(* Logix 5000 project; controller UOWHF Emulate 5570 rev 30.12; software revision 30.00; part 8 of 13 *)
(* tags used below, declared in another part *)
   UOWHF_Add_c : DINT;
   UOWHF_Msg : DINT[16];
   UOWHF_Result : DINT[16];
(* MainProgram, continued *)

   		UOWHF_Result[7]:=UOWHF_Result[7] + 421348795+UOWHF_Add_c;
   		UOWHF_Add_c.7:=UOWHF_Result[7].31;
   		UOWHF_Result[7].31:=0;
   		UOWHF_Result[8]:=UOWHF_Result[8] + 1440025142+UOWHF_Add_c;
   		UOWHF_Add_c.8:=UOWHF_Result[8].31;
   		UOWHF_Result[8].31:=0;
   	End_If;
   	If UOWHF_Msg[2].[17] Then
   		UOWHF_Result[0]:=UOWHF_Result[0] + 1919227168+UOWHF_Add_c;
   		UOWHF_Add_c.0:=UOWHF_Result[0].31;
   		UOWHF_Result[0].31:=0;
   		UOWHF_Result[1]:=UOWHF_Result[1] + 29463341+UOWHF_Add_c;
   		UOWHF_Add_c.1:=UOWHF_Result[1].31;
   		UOWHF_Result[1].31:=0;
   		UOWHF_Result[2]:=UOWHF_Result[2] + 852012451+UOWHF_Add_c;
   		UOWHF_Add_c.2:=UOWHF_Result[2].31;
   		UOWHF_Result[2].31:=0;
   		UOWHF_Result[3]:=UOWHF_Result[3] + 551239594+UOWHF_Add_c;
   		UOWHF_Add_c.3:=UOWHF_Result[3].31;
   		UOWHF_Result[3].31:=0;
   		UOWHF_Result[4]:=UOWHF_Result[4] + 213735753+UOWHF_Add_c;
   		UOWHF_Add_c.4:=UOWHF_Result[4].31;
   		UOWHF_Result[4].31:=0;
   		UOWHF_Result[5]:=UOWHF_Result[5] + 930229489+UOWHF_Add_c;
   		UOWHF_Add_c.5:=UOWHF_Result[5].31;
   		UOWHF_Result[5].31:=0;
   		UOWHF_Result[6]:=UOWHF_Result[6] + 403306511+UOWHF_Add_c;
   		UOWHF_Add_c.6:=UOWHF_Result[6].31;
   		UOWHF_Result[6].31:=0;
   		UOWHF_Result[7]:=UOWHF_Result[7] + 1320163597+UOWHF_Add_c;
   		UOWHF_Add_c.7:=UOWHF_Result[7].31;
   		UOWHF_Result[7].31:=0;
   		UOWHF_Result[8]:=UOWHF_Result[8] + 1897862563+UOWHF_Add_c;
   		UOWHF_Add_c.8:=UOWHF_Result[8].31;
   		UOWHF_Result[8].31:=0;
   	End_If;
   	If UOWHF_Msg[2].[18] Then
   		UOWHF_Result[0]:=UOWHF_Result[0] + 207957642+UOWHF_Add_c;
   		UOWHF_Add_c.0:=UOWHF_Result[0].31;
   		UOWHF_Result[0].31:=0;
   		UOWHF_Result[1]:=UOWHF_Result[1] + 1171801270+UOWHF_Add_c;
   		UOWHF_Add_c.1:=UOWHF_Result[1].31;
   		UOWHF_Result[1].31:=0;
   		UOWHF_Result[2]:=UOWHF_Result[2] + 490989868+UOWHF_Add_c;
   		UOWHF_Add_c.2:=UOWHF_Result[2].31;
   		UOWHF_Result[2].31:=0;
   		UOWHF_Result[3]:=UOWHF_Result[3] + 517478476+UOWHF_Add_c;
   		UOWHF_Add_c.3:=UOWHF_Result[3].31;
   		UOWHF_Result[3].31:=0;
   		UOWHF_Result[4]:=UOWHF_Result[4] + 709606705+UOWHF_Add_c;
   		UOWHF_Add_c.4:=UOWHF_Result[4].31;
   		UOWHF_Result[4].31:=0;
   		UOWHF_Result[5]:=UOWHF_Result[5] + 959699469+UOWHF_Add_c;
   		UOWHF_Add_c.5:=UOWHF_Result[5].31;
   		UOWHF_Result[5].31:=0;
   		UOWHF_Result[6]:=UOWHF_Result[6] + 1426433136+UOWHF_Add_c;
   		UOWHF_Add_c.6:=UOWHF_Result[6].31;
   		UOWHF_Result[6].31:=0;
   		UOWHF_Result[7]:=UOWHF_Result[7] + 861500679+UOWHF_Add_c;
   		UOWHF_Add_c.7:=UOWHF_Result[7].31;
   		UOWHF_Result[7].31:=0;
   		UOWHF_Result[8]:=UOWHF_Result[8] + 1202438537+UOWHF_Add_c;
   		UOWHF_Add_c.8:=UOWHF_Result[8].31;
   		UOWHF_Result[8].31:=0;
   	End_If;
   	If UOWHF_Msg[2].[19] Then
   		UOWHF_Result[0]:=UOWHF_Result[0] + 1004597840+UOWHF_Add_c;
   		UOWHF_Add_c.0:=UOWHF_Result[0].31;
   		UOWHF_Result[0].31:=0;
   		UOWHF_Result[1]:=UOWHF_Result[1] + 599270858+UOWHF_Add_c;
   		UOWHF_Add_c.1:=UOWHF_Result[1].31;
   		UOWHF_Result[1].31:=0;
   		UOWHF_Result[2]:=UOWHF_Result[2] + 334847739+UOWHF_Add_c;
   		UOWHF_Add_c.2:=UOWHF_Result[2].31;
   		UOWHF_Result[2].31:=0;
   		UOWHF_Result[3]:=UOWHF_Result[3] + 1969220087+UOWHF_Add_c;
   		UOWHF_Add_c.3:=UOWHF_Result[3].31;
   		UOWHF_Result[3].31:=0;
   		UOWHF_Result[4]:=UOWHF_Result[4] + 935752387+UOWHF_Add_c;
   		UOWHF_Add_c.4:=UOWHF_Result[4].31;
   		UOWHF_Result[4].31:=0;
   		UOWHF_Result[5]:=UOWHF_Result[5] + 1383478312+UOWHF_Add_c;
   		UOWHF_Add_c.5:=UOWHF_Result[5].31;
   		UOWHF_Result[5].31:=0;
   		UOWHF_Result[6]:=UOWHF_Result[6] + 138334567+UOWHF_Add_c;
   		UOWHF_Add_c.6:=UOWHF_Result[6].31;
   		UOWHF_Result[6].31:=0;
   		UOWHF_Result[7]:=UOWHF_Result[7] + 1365274530+UOWHF_Add_c;
   		UOWHF_Add_c.7:=UOWHF_Result[7].31;
   		UOWHF_Result[7].31:=0;
   		UOWHF_Result[8]:=UOWHF_Result[8] + 534270135+UOWHF_Add_c;
   		UOWHF_Add_c.8:=UOWHF_Result[8].31;
   		UOWHF_Result[8].31:=0;
   	End_If;
   	If UOWHF_Msg[2].[20] Then
   		UOWHF_Result[0]:=UOWHF_Result[0] + 638769264+UOWHF_Add_c;
   		UOWHF_Add_c.0:=UOWHF_Result[0].31;
   		UOWHF_Result[0].31:=0;
   		UOWHF_Result[1]:=UOWHF_Result[1] + 317214964+UOWHF_Add_c;
   		UOWHF_Add_c.1:=UOWHF_Result[1].31;
   		UOWHF_Result[1].31:=0;
   		UOWHF_Result[2]:=UOWHF_Result[2] + 908553039+UOWHF_Add_c;
   		UOWHF_Add_c.2:=UOWHF_Result[2].31;
   		UOWHF_Result[2].31:=0;
   		UOWHF_Result[3]:=UOWHF_Result[3] + 1054049644+UOWHF_Add_c;
   		UOWHF_Add_c.3:=UOWHF_Result[3].31;
   		UOWHF_Result[3].31:=0;
   		UOWHF_Result[4]:=UOWHF_Result[4] + 1355262167+UOWHF_Add_c;
   		UOWHF_Add_c.4:=UOWHF_Result[4].31;
   		UOWHF_Result[4].31:=0;
   		UOWHF_Result[5]:=UOWHF_Result[5] + 1333398518+UOWHF_Add_c;
   		UOWHF_Add_c.5:=UOWHF_Result[5].31;
   		UOWHF_Result[5].31:=0;
   		UOWHF_Result[6]:=UOWHF_Result[6] + 923137105+UOWHF_Add_c;
   		UOWHF_Add_c.6:=UOWHF_Result[6].31;
   		UOWHF_Result[6].31:=0;
   		UOWHF_Result[7]:=UOWHF_Result[7] + 1603787279+UOWHF_Add_c;
   		UOWHF_Add_c.7:=UOWHF_Result[7].31;
   		UOWHF_Result[7].31:=0;
   		UOWHF_Result[8]:=UOWHF_Result[8] + 215241896+UOWHF_Add_c;
   		UOWHF_Add_c.8:=UOWHF_Result[8].31;
   		UOWHF_Result[8].31:=0;
   	End_If;
   	If UOWHF_Msg[2].[21] Then
   		UOWHF_Result[0]:=UOWHF_Result[0] + 1253585795+UOWHF_Add_c;
   		UOWHF_Add_c.0:=UOWHF_Result[0].31;
   		UOWHF_Result[0].31:=0;
   		UOWHF_Result[1]:=UOWHF_Result[1] + 1774567950+UOWHF_Add_c;
   		UOWHF_Add_c.1:=UOWHF_Result[1].31;
   		UOWHF_Result[1].31:=0;
   		UOWHF_Result[2]:=UOWHF_Result[2] + 1348389163+UOWHF_Add_c;
   		UOWHF_Add_c.2:=UOWHF_Result[2].31;
   		UOWHF_Result[2].31:=0;
   		UOWHF_Result[3]:=UOWHF_Result[3] + 1776776512+UOWHF_Add_c;
   		UOWHF_Add_c.3:=UOWHF_Result[3].31;
   		UOWHF_Result[3].31:=0;
   		UOWHF_Result[4]:=UOWHF_Result[4] + 1887727344+UOWHF_Add_c;
   		UOWHF_Add_c.4:=UOWHF_Result[4].31;
   		UOWHF_Result[4].31:=0;
   		UOWHF_Result[5]:=UOWHF_Result[5] + 420280741+UOWHF_Add_c;
   		UOWHF_Add_c.5:=UOWHF_Result[5].31;
   		UOWHF_Result[5].31:=0;
   		UOWHF_Result[6]:=UOWHF_Result[6] + 1390579328+UOWHF_Add_c;
   		UOWHF_Add_c.6:=UOWHF_Result[6].31;
   		UOWHF_Result[6].31:=0;
   		UOWHF_Result[7]:=UOWHF_Result[7] + 928509381+UOWHF_Add_c;
   		UOWHF_Add_c.7:=UOWHF_Result[7].31;
   		UOWHF_Result[7].31:=0;
   		UOWHF_Result[8]:=UOWHF_Result[8] + 1507051281+UOWHF_Add_c;
   		UOWHF_Add_c.8:=UOWHF_Result[8].31;
   		UOWHF_Result[8].31:=0;
   	End_If;
   	If UOWHF_Msg[2].[22] Then
   		UOWHF_Result[0]:=UOWHF_Result[0] + 1291966163+UOWHF_Add_c;
   		UOWHF_Add_c.0:=UOWHF_Result[0].31;
   		UOWHF_Result[0].31:=0;
   		UOWHF_Result[1]:=UOWHF_Result[1] + 466028181+UOWHF_Add_c;
   		UOWHF_Add_c.1:=UOWHF_Result[1].31;
   		UOWHF_Result[1].31:=0;
   		UOWHF_Result[2]:=UOWHF_Result[2] + 1269422310+UOWHF_Add_c;
   		UOWHF_Add_c.2:=UOWHF_Result[2].31;
   		UOWHF_Result[2].31:=0;
   		UOWHF_Result[3]:=UOWHF_Result[3] + 167272220+UOWHF_Add_c;
   		UOWHF_Add_c.3:=UOWHF_Result[3].31;
   		UOWHF_Result[3].31:=0;
   		UOWHF_Result[4]:=UOWHF_Result[4] + 1812138151+UOWHF_Add_c;
   		UOWHF_Add_c.4:=UOWHF_Result[4].31;
   		UOWHF_Result[4].31:=0;
   		UOWHF_Result[5]:=UOWHF_Result[5] + 2028840979+UOWHF_Add_c;
   		UOWHF_Add_c.5:=UOWHF_Result[5].31;
   		UOWHF_Result[5].31:=0;
   		UOWHF_Result[6]:=UOWHF_Result[6] + 1588214460+UOWHF_Add_c;
   		UOWHF_Add_c.6:=UOWHF_Result[6].31;
   		UOWHF_Result[6].31:=0;
   		UOWHF_Result[7]:=UOWHF_Result[7] + 1912044568+UOWHF_Add_c;
   		UOWHF_Add_c.7:=UOWHF_Result[7].31;
   		UOWHF_Result[7].31:=0;
   		UOWHF_Result[8]:=UOWHF_Result[8] + 690703953+UOWHF_Add_c;
   		UOWHF_Add_c.8:=UOWHF_Result[8].31;
   		UOWHF_Result[8].31:=0;
   	End_If;
   	If UOWHF_Msg[2].[23] Then
   		UOWHF_Result[0]:=UOWHF_Result[0] + 1665444751+UOWHF_Add_c;
   		UOWHF_Add_c.0:=UOWHF_Result[0].31;
   		UOWHF_Result[0].31:=0;
   		UOWHF_Result[1]:=UOWHF_Result[1] + 878466108+UOWHF_Add_c;
   		UOWHF_Add_c.1:=UOWHF_Result[1].31;
   		UOWHF_Result[1].31:=0;
   		UOWHF_Result[2]:=UOWHF_Result[2] + 1084953660+UOWHF_Add_c;
   		UOWHF_Add_c.2:=UOWHF_Result[2].31;
   		UOWHF_Result[2].31:=0;
   		UOWHF_Result[3]:=UOWHF_Result[3] + 1182760719+UOWHF_Add_c;
   		UOWHF_Add_c.3:=UOWHF_Result[3].31;
   		UOWHF_Result[3].31:=0;
   		UOWHF_Result[4]:=UOWHF_Result[4] + 1329395022+UOWHF_Add_c;
   		UOWHF_Add_c.4:=UOWHF_Result[4].31;
   		UOWHF_Result[4].31:=0;
   		UOWHF_Result[5]:=UOWHF_Result[5] + 2000087125+UOWHF_Add_c;
   		UOWHF_Add_c.5:=UOWHF_Result[5].31;
   		UOWHF_Result[5].31:=0;
   		UOWHF_Result[6]:=UOWHF_Result[6] + 1154519389+UOWHF_Add_c;
   		UOWHF_Add_c.6:=UOWHF_Result[6].31;
   		UOWHF_Result[6].31:=0;
   		UOWHF_Result[7]:=UOWHF_Result[7] + 301344254+UOWHF_Add_c;
   		UOWHF_Add_c.7:=UOWHF_Result[7].31;
   		UOWHF_Result[7].31:=0;
   		UOWHF_Result[8]:=UOWHF_Result[8] + 1297674993+UOWHF_Add_c;
   		UOWHF_Add_c.8:=UOWHF_Result[8].31;
   		UOWHF_Result[8].31:=0;
   	End_If;
   	If UOWHF_Msg[2].[24] Then
   		UOWHF_Result[0]:=UOWHF_Result[0] + 558242359+UOWHF_Add_c;
   		UOWHF_Add_c.0:=UOWHF_Result[0].31;
   		UOWHF_Result[0].31:=0;
   		UOWHF_Result[1]:=UOWHF_Result[1] + 959605875+UOWHF_Add_c;
   		UOWHF_Add_c.1:=UOWHF_Result[1].31;
   		UOWHF_Result[1].31:=0;
   		UOWHF_Result[2]:=UOWHF_Result[2] + 1409764266+UOWHF_Add_c;
   		UOWHF_Add_c.2:=UOWHF_Result[2].31;
   		UOWHF_Result[2].31:=0;
   		UOWHF_Result[3]:=UOWHF_Result[3] + 1619308583+UOWHF_Add_c;
   		UOWHF_Add_c.3:=UOWHF_Result[3].31;
   		UOWHF_Result[3].31:=0;
   		UOWHF_Result[4]:=UOWHF_Result[4] + 642811496+UOWHF_Add_c;
   		UOWHF_Add_c.4:=UOWHF_Result[4].31;
   		UOWHF_Result[4].31:=0;
   		UOWHF_Result[5]:=UOWHF_Result[5] + 1911637828+UOWHF_Add_c;
   		UOWHF_Add_c.5:=UOWHF_Result[5].31;
   		UOWHF_Result[5].31:=0;
   		UOWHF_Result[6]:=UOWHF_Result[6] + 688982836+UOWHF_Add_c;
   		UOWHF_Add_c.6:=UOWHF_Result[6].31;
   		UOWHF_Result[6].31:=0;
   		UOWHF_Result[7]:=UOWHF_Result[7] + 189891926+UOWHF_Add_c;
   		UOWHF_Add_c.7:=UOWHF_Result[7].31;
   		UOWHF_Result[7].31:=0;
   		UOWHF_Result[8]:=UOWHF_Result[8] + 1047838333+UOWHF_Add_c;
   		UOWHF_Add_c.8:=UOWHF_Result[8].31;
   		UOWHF_Result[8].31:=0;
   	End_If;
   	If UOWHF_Msg[2].[25] Then
   		UOWHF_Result[0]:=UOWHF_Result[0] + 166408324+UOWHF_Add_c;
   		UOWHF_Add_c.0:=UOWHF_Result[0].31;
   		UOWHF_Result[0].31:=0;
   		UOWHF_Result[1]:=UOWHF_Result[1] + 1090081190+UOWHF_Add_c;
   		UOWHF_Add_c.1:=UOWHF_Result[1].31;
   		UOWHF_Result[1].31:=0;
   		UOWHF_Result[2]:=UOWHF_Result[2] + 1222902067+UOWHF_Add_c;
   		UOWHF_Add_c.2:=UOWHF_Result[2].31;
   		UOWHF_Result[2].31:=0;
   		UOWHF_Result[3]:=UOWHF_Result[3] + 740886112+UOWHF_Add_c;
   		UOWHF_Add_c.3:=UOWHF_Result[3].31;
   		UOWHF_Result[3].31:=0;
   		UOWHF_Result[4]:=UOWHF_Result[4] + 963550939+UOWHF_Add_c;
   		UOWHF_Add_c.4:=UOWHF_Result[4].31;
   		UOWHF_Result[4].31:=0;
   		UOWHF_Result[5]:=UOWHF_Result[5] + 965997722+UOWHF_Add_c;
   		UOWHF_Add_c.5:=UOWHF_Result[5].31;
   		UOWHF_Result[5].31:=0;
   		UOWHF_Result[6]:=UOWHF_Result[6] + 1814719293+UOWHF_Add_c;
   		UOWHF_Add_c.6:=UOWHF_Result[6].31;
   		UOWHF_Result[6].31:=0;
   		UOWHF_Result[7]:=UOWHF_Result[7] + 942657862+UOWHF_Add_c;
   		UOWHF_Add_c.7:=UOWHF_Result[7].31;
   		UOWHF_Result[7].31:=0;
   		UOWHF_Result[8]:=UOWHF_Result[8] + 1993997569+UOWHF_Add_c;
   		UOWHF_Add_c.8:=UOWHF_Result[8].31;
   		UOWHF_Result[8].31:=0;
   	End_If;
   	If UOWHF_Msg[2].[26] Then
   		UOWHF_Result[0]:=UOWHF_Result[0] + 63286127+UOWHF_Add_c;
   		UOWHF_Add_c.0:=UOWHF_Result[0].31;
   		UOWHF_Result[0].31:=0;
   		UOWHF_Result[1]:=UOWHF_Result[1] + 99678506+UOWHF_Add_c;
   		UOWHF_Add_c.1:=UOWHF_Result[1].31;
   		UOWHF_Result[1].31:=0;
   		UOWHF_Result[2]:=UOWHF_Result[2] + 323238799+UOWHF_Add_c;
   		UOWHF_Add_c.2:=UOWHF_Result[2].31;
   		UOWHF_Result[2].31:=0;
   		UOWHF_Result[3]:=UOWHF_Result[3] + 1161946555+UOWHF_Add_c;
   		UOWHF_Add_c.3:=UOWHF_Result[3].31;
   		UOWHF_Result[3].31:=0;
   		UOWHF_Result[4]:=UOWHF_Result[4] + 444321833+UOWHF_Add_c;
   		UOWHF_Add_c.4:=UOWHF_Result[4].31;
   		UOWHF_Result[4].31:=0;
   		UOWHF_Result[5]:=UOWHF_Result[5] + 1552943728+UOWHF_Add_c;
   		UOWHF_Add_c.5:=UOWHF_Result[5].31;
   		UOWHF_Result[5].31:=0;
   		UOWHF_Result[6]:=UOWHF_Result[6] + 1367212046+UOWHF_Add_c;
   		UOWHF_Add_c.6:=UOWHF_Result[6].31;
   		UOWHF_Result[6].31:=0;
   		UOWHF_Result[7]:=UOWHF_Result[7] + 1197605653+UOWHF_Add_c;
   		UOWHF_Add_c.7:=UOWHF_Result[7].31;
   		UOWHF_Result[7].31:=0;
   		UOWHF_Result[8]:=UOWHF_Result[8] + 473086606+UOWHF_Add_c;
   		UOWHF_Add_c.8:=UOWHF_Result[8].31;
   		UOWHF_Result[8].31:=0;
   	End_If;
   	If UOWHF_Msg[2].[27] Then
   		UOWHF_Result[0]:=UOWHF_Result[0] + 1220273658+UOWHF_Add_c;
   		UOWHF_Add_c.0:=UOWHF_Result[0].31;
   		UOWHF_Result[0].31:=0;
   		UOWHF_Result[1]:=UOWHF_Result[1] + 2138805728+UOWHF_Add_c;
   		UOWHF_Add_c.1:=UOWHF_Result[1].31;
   		UOWHF_Result[1].31:=0;
   		UOWHF_Result[2]:=UOWHF_Result[2] + 105977955+UOWHF_Add_c;
   		UOWHF_Add_c.2:=UOWHF_Result[2].31;
   		UOWHF_Result[2].31:=0;
   		UOWHF_Result[3]:=UOWHF_Result[3] + 848247904+UOWHF_Add_c;
   		UOWHF_Add_c.3:=UOWHF_Result[3].31;
   		UOWHF_Result[3].31:=0;
   		UOWHF_Result[4]:=UOWHF_Result[4] + 105843336+UOWHF_Add_c;
   		UOWHF_Add_c.4:=UOWHF_Result[4].31;
   		UOWHF_Result[4].31:=0;
   		UOWHF_Result[5]:=UOWHF_Result[5] + 1286591821+UOWHF_Add_c;
   		UOWHF_Add_c.5:=UOWHF_Result[5].31;
   		UOWHF_Result[5].31:=0;
   		UOWHF_Result[6]:=UOWHF_Result[6] + 155040163+UOWHF_Add_c;
   		UOWHF_Add_c.6:=UOWHF_Result[6].31;
   		UOWHF_Result[6].31:=0;
   		UOWHF_Result[7]:=UOWHF_Result[7] + 1480293425+UOWHF_Add_c;
   		UOWHF_Add_c.7:=UOWHF_Result[7].31;
   		UOWHF_Result[7].31:=0;
   		UOWHF_Result[8]:=UOWHF_Result[8] + 1440769872+UOWHF_Add_c;
   		UOWHF_Add_c.8:=UOWHF_Result[8].31;
   		UOWHF_Result[8].31:=0;
   	End_If;
   	If UOWHF_Msg[2].[28] Then
   		UOWHF_Result[0]:=UOWHF_Result[0] + 1372096306+UOWHF_Add_c;
   		UOWHF_Add_c.0:=UOWHF_Result[0].31;
   		UOWHF_Result[0].31:=0;
   		UOWHF_Result[1]:=UOWHF_Result[1] + 507063276+UOWHF_Add_c;
   		UOWHF_Add_c.1:=UOWHF_Result[1].31;
   		UOWHF_Result[1].31:=0;
   		UOWHF_Result[2]:=UOWHF_Result[2] + 1427839543+UOWHF_Add_c;
   		UOWHF_Add_c.2:=UOWHF_Result[2].31;
   		UOWHF_Result[2].31:=0;
   		UOWHF_Result[3]:=UOWHF_Result[3] + 1125336766+UOWHF_Add_c;
   		UOWHF_Add_c.3:=UOWHF_Result[3].31;
   		UOWHF_Result[3].31:=0;
   		UOWHF_Result[4]:=UOWHF_Result[4] + 999982338+UOWHF_Add_c;
   		UOWHF_Add_c.4:=UOWHF_Result[4].31;
   		UOWHF_Result[4].31:=0;
   		UOWHF_Result[5]:=UOWHF_Result[5] + 1914412456+UOWHF_Add_c;
   		UOWHF_Add_c.5:=UOWHF_Result[5].31;
   		UOWHF_Result[5].31:=0;
   		UOWHF_Result[6]:=UOWHF_Result[6] + 974480105+UOWHF_Add_c;
   		UOWHF_Add_c.6:=UOWHF_Result[6].31;
   		UOWHF_Result[6].31:=0;
   		UOWHF_Result[7]:=UOWHF_Result[7] + 1780395916+UOWHF_Add_c;
   		UOWHF_Add_c.7:=UOWHF_Result[7].31;
   		UOWHF_Result[7].31:=0;
   		UOWHF_Result[8]:=UOWHF_Result[8] + 33420938+UOWHF_Add_c;
   		UOWHF_Add_c.8:=UOWHF_Result[8].31;
   		UOWHF_Result[8].31:=0;
   	End_If;
   	If UOWHF_Msg[2].[29] Then
   		UOWHF_Result[0]:=UOWHF_Result[0] + 976400534+UOWHF_Add_c;
   		UOWHF_Add_c.0:=UOWHF_Result[0].31;
   		UOWHF_Result[0].31:=0;
   		UOWHF_Result[1]:=UOWHF_Result[1] + 1662471994+UOWHF_Add_c;
   		UOWHF_Add_c.1:=UOWHF_Result[1].31;
   		UOWHF_Result[1].31:=0;
   		UOWHF_Result[2]:=UOWHF_Result[2] + 772226603+UOWHF_Add_c;
   		UOWHF_Add_c.2:=UOWHF_Result[2].31;
   		UOWHF_Result[2].31:=0;
   		UOWHF_Result[3]:=UOWHF_Result[3] + 1441513688+UOWHF_Add_c;
   		UOWHF_Add_c.3:=UOWHF_Result[3].31;
   		UOWHF_Result[3].31:=0;
   		UOWHF_Result[4]:=UOWHF_Result[4] + 1888957472+UOWHF_Add_c;
   		UOWHF_Add_c.4:=UOWHF_Result[4].31;
   		UOWHF_Result[4].31:=0;
   		UOWHF_Result[5]:=UOWHF_Result[5] + 483859248+UOWHF_Add_c;
   		UOWHF_Add_c.5:=UOWHF_Result[5].31;
   		UOWHF_Result[5].31:=0;
   		UOWHF_Result[6]:=UOWHF_Result[6] + 822038845+UOWHF_Add_c;
   		UOWHF_Add_c.6:=UOWHF_Result[6].31;
   		UOWHF_Result[6].31:=0;
   		UOWHF_Result[7]:=UOWHF_Result[7] + 1422074512+UOWHF_Add_c;
   		UOWHF_Add_c.7:=UOWHF_Result[7].31;
   		UOWHF_Result[7].31:=0;
   		UOWHF_Result[8]:=UOWHF_Result[8] + 1027247335+UOWHF_Add_c;
   		UOWHF_Add_c.8:=UOWHF_Result[8].31;
   		UOWHF_Result[8].31:=0;
   	End_If;
   	If UOWHF_Msg[2].[30] Then
   		UOWHF_Result[0]:=UOWHF_Result[0] + 1714194303+UOWHF_Add_c;
   		UOWHF_Add_c.0:=UOWHF_Result[0].31;
   		UOWHF_Result[0].31:=0;
   		UOWHF_Result[1]:=UOWHF_Result[1] + 2010412813+UOWHF_Add_c;
   		UOWHF_Add_c.1:=UOWHF_Result[1].31;
   		UOWHF_Result[1].31:=0;
   		UOWHF_Result[2]:=UOWHF_Result[2] + 312944695+UOWHF_Add_c;
   		UOWHF_Add_c.2:=UOWHF_Result[2].31;
   		UOWHF_Result[2].31:=0;
   		UOWHF_Result[3]:=UOWHF_Result[3] + 520236415+UOWHF_Add_c;
   		UOWHF_Add_c.3:=UOWHF_Result[3].31;
   		UOWHF_Result[3].31:=0;
   		UOWHF_Result[4]:=UOWHF_Result[4] + 667902072+UOWHF_Add_c;
   		UOWHF_Add_c.4:=UOWHF_Result[4].31;
   		UOWHF_Result[4].31:=0;
   		UOWHF_Result[5]:=UOWHF_Result[5] + 1787858584+UOWHF_Add_c;
   		UOWHF_Add_c.5:=UOWHF_Result[5].31;
   		UOWHF_Result[5].31:=0;
   		UOWHF_Result[6]:=UOWHF_Result[6] + 1416792661+UOWHF_Add_c;
   		UOWHF_Add_c.6:=UOWHF_Result[6].31;
   		UOWHF_Result[6].31:=0;
   		UOWHF_Result[7]:=UOWHF_Result[7] + 1986385854+UOWHF_Add_c;
   		UOWHF_Add_c.7:=UOWHF_Result[7].31;
   		UOWHF_Result[7].31:=0;
   		UOWHF_Result[8]:=UOWHF_Result[8] + 80966913+UOWHF_Add_c;
   		UOWHF_Add_c.8:=UOWHF_Result[8].31;
   		UOWHF_Result[8].31:=0;
   	End_If;
   	If UOWHF_Msg[2].[31] Then
   		UOWHF_Result[0]:=UOWHF_Result[0] + 142019018+UOWHF_Add_c;
   		UOWHF_Add_c.0:=UOWHF_Result[0].31;
   		UOWHF_Result[0].31:=0;
   		UOWHF_Result[1]:=UOWHF_Result[1] + 1347023134+UOWHF_Add_c;
   		UOWHF_Add_c.1:=UOWHF_Result[1].31;
   		UOWHF_Result[1].31:=0;
   		UOWHF_Result[2]:=UOWHF_Result[2] + 323000754+UOWHF_Add_c;
   		UOWHF_Add_c.2:=UOWHF_Result[2].31;
   		UOWHF_Result[2].31:=0;
   		UOWHF_Result[3]:=UOWHF_Result[3] + 1411034496+UOWHF_Add_c;
   		UOWHF_Add_c.3:=UOWHF_Result[3].31;
   		UOWHF_Result[3].31:=0;
   		UOWHF_Result[4]:=UOWHF_Result[4] + 1353462926+UOWHF_Add_c;
   		UOWHF_Add_c.4:=UOWHF_Result[4].31;
   		UOWHF_Result[4].31:=0;
   		UOWHF_Result[5]:=UOWHF_Result[5] + 885192095+UOWHF_Add_c;
   		UOWHF_Add_c.5:=UOWHF_Result[5].31;
   		UOWHF_Result[5].31:=0;
   		UOWHF_Result[6]:=UOWHF_Result[6] + 101022159+UOWHF_Add_c;
   		UOWHF_Add_c.6:=UOWHF_Result[6].31;
   		UOWHF_Result[6].31:=0;
   		UOWHF_Result[7]:=UOWHF_Result[7] + 1892280229+UOWHF_Add_c;
   		UOWHF_Add_c.7:=UOWHF_Result[7].31;
   		UOWHF_Result[7].31:=0;
   		UOWHF_Result[8]:=UOWHF_Result[8] + 165464048+UOWHF_Add_c;
   		UOWHF_Add_c.8:=UOWHF_Result[8].31;
   		UOWHF_Result[8].31:=0;
   	End_If;
   	If UOWHF_Msg[3].[0] Then
   		UOWHF_Result[0]:=UOWHF_Result[0] + 404019456+UOWHF_Add_c;
   		UOWHF_Add_c.0:=UOWHF_Result[0].31;
   		UOWHF_Result[0].31:=0;
   		UOWHF_Result[1]:=UOWHF_Result[1] + 1191571511+UOWHF_Add_c;
   		UOWHF_Add_c.1:=UOWHF_Result[1].31;
   		UOWHF_Result[1].31:=0;
   		UOWHF_Result[2]:=UOWHF_Result[2] + 744168101+UOWHF_Add_c;
   		UOWHF_Add_c.2:=UOWHF_Result[2].31;
   		UOWHF_Result[2].31:=0;
   		UOWHF_Result[3]:=UOWHF_Result[3] + 822803911+UOWHF_Add_c;
   		UOWHF_Add_c.3:=UOWHF_Result[3].31;
   		UOWHF_Result[3].31:=0;
   		UOWHF_Result[4]:=UOWHF_Result[4] + 1922930597+UOWHF_Add_c;
   		UOWHF_Add_c.4:=UOWHF_Result[4].31;
   		UOWHF_Result[4].31:=0;
   		UOWHF_Result[5]:=UOWHF_Result[5] + 1557038461+UOWHF_Add_c;
   		UOWHF_Add_c.5:=UOWHF_Result[5].31;
   		UOWHF_Result[5].31:=0;
   		UOWHF_Result[6]:=UOWHF_Result[6] + 1297088610+UOWHF_Add_c;
   		UOWHF_Add_c.6:=UOWHF_Result[6].31;
   		UOWHF_Result[6].31:=0;
   		UOWHF_Result[7]:=UOWHF_Result[7] + 1640767354+UOWHF_Add_c;
   		UOWHF_Add_c.7:=UOWHF_Result[7].31;
   		UOWHF_Result[7].31:=0;
   		UOWHF_Result[8]:=UOWHF_Result[8] + 564595313+UOWHF_Add_c;
   		UOWHF_Add_c.8:=UOWHF_Result[8].31;
   		UOWHF_Result[8].31:=0;
   	End_If;
   	If UOWHF_Msg[3].[1] Then
   		UOWHF_Result[0]:=UOWHF_Result[0] + 1300701096+UOWHF_Add_c;
   		UOWHF_Add_c.0:=UOWHF_Result[0].31;
   		UOWHF_Result[0].31:=0;
   		UOWHF_Result[1]:=UOWHF_Result[1] + 740702294+UOWHF_Add_c;
   		UOWHF_Add_c.1:=UOWHF_Result[1].31;
   		UOWHF_Result[1].31:=0;
   		UOWHF_Result[2]:=UOWHF_Result[2] + 69145646+UOWHF_Add_c;
   		UOWHF_Add_c.2:=UOWHF_Result[2].31;
   		UOWHF_Result[2].31:=0;
   		UOWHF_Result[3]:=UOWHF_Result[3] + 1305021096+UOWHF_Add_c;
   		UOWHF_Add_c.3:=UOWHF_Result[3].31;
   		UOWHF_Result[3].31:=0;
   		UOWHF_Result[4]:=UOWHF_Result[4] + 1394686303+UOWHF_Add_c;
   		UOWHF_Add_c.4:=UOWHF_Result[4].31;
   		UOWHF_Result[4].31:=0;
   		UOWHF_Result[5]:=UOWHF_Result[5] + 867008968+UOWHF_Add_c;
   		UOWHF_Add_c.5:=UOWHF_Result[5].31;
   		UOWHF_Result[5].31:=0;
   		UOWHF_Result[6]:=UOWHF_Result[6] + 1159266556+UOWHF_Add_c;
   		UOWHF_Add_c.6:=UOWHF_Result[6].31;
   		UOWHF_Result[6].31:=0;
   		UOWHF_Result[7]:=UOWHF_Result[7] + 127314732+UOWHF_Add_c;
   		UOWHF_Add_c.7:=UOWHF_Result[7].31;
   		UOWHF_Result[7].31:=0;
   		UOWHF_Result[8]:=UOWHF_Result[8] + 537818420+UOWHF_Add_c;
   		UOWHF_Add_c.8:=UOWHF_Result[8].31;
   		UOWHF_Result[8].31:=0;
   	End_If;
   	If UOWHF_Msg[3].[2] Then
   		UOWHF_Result[0]:=UOWHF_Result[0] + 686229662+UOWHF_Add_c;
   		UOWHF_Add_c.0:=UOWHF_Result[0].31;
   		UOWHF_Result[0].31:=0;
   		UOWHF_Result[1]:=UOWHF_Result[1] + 519859819+UOWHF_Add_c;
   		UOWHF_Add_c.1:=UOWHF_Result[1].31;
   		UOWHF_Result[1].31:=0;
   		UOWHF_Result[2]:=UOWHF_Result[2] + 1370828025+UOWHF_Add_c;
   		UOWHF_Add_c.2:=UOWHF_Result[2].31;
   		UOWHF_Result[2].31:=0;
   		UOWHF_Result[3]:=UOWHF_Result[3] + 2030093876+UOWHF_Add_c;
   		UOWHF_Add_c.3:=UOWHF_Result[3].31;
   		UOWHF_Result[3].31:=0;
   		UOWHF_Result[4]:=UOWHF_Result[4] + 912557543+UOWHF_Add_c;
   		UOWHF_Add_c.4:=UOWHF_Result[4].31;
   		UOWHF_Result[4].31:=0;
   		UOWHF_Result[5]:=UOWHF_Result[5] + 1074494947+UOWHF_Add_c;
   		UOWHF_Add_c.5:=UOWHF_Result[5].31;
   		UOWHF_Result[5].31:=0;
   		UOWHF_Result[6]:=UOWHF_Result[6] + 962454511+UOWHF_Add_c;
   		UOWHF_Add_c.6:=UOWHF_Result[6].31;
   		UOWHF_Result[6].31:=0;
   		UOWHF_Result[7]:=UOWHF_Result[7] + 717388161+UOWHF_Add_c;
   		UOWHF_Add_c.7:=UOWHF_Result[7].31;
   		UOWHF_Result[7].31:=0;
   		UOWHF_Result[8]:=UOWHF_Result[8] + 1855883681+UOWHF_Add_c;
   		UOWHF_Add_c.8:=UOWHF_Result[8].31;
   		UOWHF_Result[8].31:=0;
   	End_If;
   	If UOWHF_Msg[3].[3] Then
   		UOWHF_Result[0]:=UOWHF_Result[0] + 81890441+UOWHF_Add_c;
   		UOWHF_Add_c.0:=UOWHF_Result[0].31;
   		UOWHF_Result[0].31:=0;
   		UOWHF_Result[1]:=UOWHF_Result[1] + 1611695652+UOWHF_Add_c;
   		UOWHF_Add_c.1:=UOWHF_Result[1].31;
   		UOWHF_Result[1].31:=0;
   		UOWHF_Result[2]:=UOWHF_Result[2] + 459192051+UOWHF_Add_c;
   		UOWHF_Add_c.2:=UOWHF_Result[2].31;
   		UOWHF_Result[2].31:=0;
   		UOWHF_Result[3]:=UOWHF_Result[3] + 1560790570+UOWHF_Add_c;
   		UOWHF_Add_c.3:=UOWHF_Result[3].31;
   		UOWHF_Result[3].31:=0;
   		UOWHF_Result[4]:=UOWHF_Result[4] + 1332180995+UOWHF_Add_c;
   		UOWHF_Add_c.4:=UOWHF_Result[4].31;
   		UOWHF_Result[4].31:=0;
   		UOWHF_Result[5]:=UOWHF_Result[5] + 1745313226+UOWHF_Add_c;
   		UOWHF_Add_c.5:=UOWHF_Result[5].31;
   		UOWHF_Result[5].31:=0;
   		UOWHF_Result[6]:=UOWHF_Result[6] + 1483887170+UOWHF_Add_c;
   		UOWHF_Add_c.6:=UOWHF_Result[6].31;
   		UOWHF_Result[6].31:=0;
   		UOWHF_Result[7]:=UOWHF_Result[7] + 767952137+UOWHF_Add_c;
   		UOWHF_Add_c.7:=UOWHF_Result[7].31;
   		UOWHF_Result[7].31:=0;
   		UOWHF_Result[8]:=UOWHF_Result[8] + 1769752883+UOWHF_Add_c;
   		UOWHF_Add_c.8:=UOWHF_Result[8].31;
   		UOWHF_Result[8].31:=0;
   	End_If;
   	If UOWHF_Msg[3].[4] Then
   		UOWHF_Result[0]:=UOWHF_Result[0] + 2037848486+UOWHF_Add_c;
   		UOWHF_Add_c.0:=UOWHF_Result[0].31;
   		UOWHF_Result[0].31:=0;
   		UOWHF_Result[1]:=UOWHF_Result[1] + 1759404806+UOWHF_Add_c;
   		UOWHF_Add_c.1:=UOWHF_Result[1].31;
   		UOWHF_Result[1].31:=0;
   		UOWHF_Result[2]:=UOWHF_Result[2] + 1391748728+UOWHF_Add_c;
   		UOWHF_Add_c.2:=UOWHF_Result[2].31;
   		UOWHF_Result[2].31:=0;
   		UOWHF_Result[3]:=UOWHF_Result[3] + 1205400143+UOWHF_Add_c;
   		UOWHF_Add_c.3:=UOWHF_Result[3].31;
   		UOWHF_Result[3].31:=0;
   		UOWHF_Result[4]:=UOWHF_Result[4] + 547556167+UOWHF_Add_c;
   		UOWHF_Add_c.4:=UOWHF_Result[4].31;
   		UOWHF_Result[4].31:=0;
   		UOWHF_Result[5]:=UOWHF_Result[5] + 2035664608+UOWHF_Add_c;
   		UOWHF_Add_c.5:=UOWHF_Result[5].31;
   		UOWHF_Result[5].31:=0;
   		UOWHF_Result[6]:=UOWHF_Result[6] + 1559257416+UOWHF_Add_c;
   		UOWHF_Add_c.6:=UOWHF_Result[6].31;
   		UOWHF_Result[6].31:=0;
   		UOWHF_Result[7]:=UOWHF_Result[7] + 870549215+UOWHF_Add_c;
   		UOWHF_Add_c.7:=UOWHF_Result[7].31;
   		UOWHF_Result[7].31:=0;
   		UOWHF_Result[8]:=UOWHF_Result[8] + 539229582+UOWHF_Add_c;
   		UOWHF_Add_c.8:=UOWHF_Result[8].31;
   		UOWHF_Result[8].31:=0;
   	End_If;
   	If UOWHF_Msg[3].[5] Then
   		UOWHF_Result[0]:=UOWHF_Result[0] + 1501452002+UOWHF_Add_c;
   		UOWHF_Add_c.0:=UOWHF_Result[0].31;
   		UOWHF_Result[0].31:=0;
   		UOWHF_Result[1]:=UOWHF_Result[1] + 1244431443+UOWHF_Add_c;
   		UOWHF_Add_c.1:=UOWHF_Result[1].31;
   		UOWHF_Result[1].31:=0;
   		UOWHF_Result[2]:=UOWHF_Result[2] + 1313958277+UOWHF_Add_c;
   		UOWHF_Add_c.2:=UOWHF_Result[2].31;
   		UOWHF_Result[2].31:=0;
   		UOWHF_Result[3]:=UOWHF_Result[3] + 712802192+UOWHF_Add_c;
   		UOWHF_Add_c.3:=UOWHF_Result[3].31;
   		UOWHF_Result[3].31:=0;
   		UOWHF_Result[4]:=UOWHF_Result[4] + 2081310582+UOWHF_Add_c;
   		UOWHF_Add_c.4:=UOWHF_Result[4].31;
   		UOWHF_Result[4].31:=0;
   		UOWHF_Result[5]:=UOWHF_Result[5] + 32566088+UOWHF_Add_c;
   		UOWHF_Add_c.5:=UOWHF_Result[5].31;
   		UOWHF_Result[5].31:=0;
   		UOWHF_Result[6]:=UOWHF_Result[6] + 2064972158+UOWHF_Add_c;
   		UOWHF_Add_c.6:=UOWHF_Result[6].31;
   		UOWHF_Result[6].31:=0;
   		UOWHF_Result[7]:=UOWHF_Result[7] + 650601391+UOWHF_Add_c;
   		UOWHF_Add_c.7:=UOWHF_Result[7].31;
   		UOWHF_Result[7].31:=0;
   		UOWHF_Result[8]:=UOWHF_Result[8] + 1456400780+UOWHF_Add_c;
   		UOWHF_Add_c.8:=UOWHF_Result[8].31;
   		UOWHF_Result[8].31:=0;
   	End_If;
   	If UOWHF_Msg[3].[6] Then
   		UOWHF_Result[0]:=UOWHF_Result[0] + 617501499+UOWHF_Add_c;
   		UOWHF_Add_c.0:=UOWHF_Result[0].31;
   		UOWHF_Result[0].31:=0;
   		UOWHF_Result[1]:=UOWHF_Result[1] + 1754016077+UOWHF_Add_c;
   		UOWHF_Add_c.1:=UOWHF_Result[1].31;
   		UOWHF_Result[1].31:=0;
   		UOWHF_Result[2]:=UOWHF_Result[2] + 2029585615+UOWHF_Add_c;
   		UOWHF_Add_c.2:=UOWHF_Result[2].31;
   		UOWHF_Result[2].31:=0;
   		UOWHF_Result[3]:=UOWHF_Result[3] + 355961793+UOWHF_Add_c;
   		UOWHF_Add_c.3:=UOWHF_Result[3].31;
   		UOWHF_Result[3].31:=0;
   		UOWHF_Result[4]:=UOWHF_Result[4] + 235264645+UOWHF_Add_c;
   		UOWHF_Add_c.4:=UOWHF_Result[4].31;
   		UOWHF_Result[4].31:=0;
   		UOWHF_Result[5]:=UOWHF_Result[5] + 1625867090+UOWHF_Add_c;
   		UOWHF_Add_c.5:=UOWHF_Result[5].31;
   		UOWHF_Result[5].31:=0;
   		UOWHF_Result[6]:=UOWHF_Result[6] + 1929512258+UOWHF_Add_c;
   		UOWHF_Add_c.6:=UOWHF_Result[6].31;
   		UOWHF_Result[6].31:=0;
   		UOWHF_Result[7]:=UOWHF_Result[7] + 274890974+UOWHF_Add_c;
   		UOWHF_Add_c.7:=UOWHF_Result[7].31;
   		UOWHF_Result[7].31:=0;
   		UOWHF_Result[8]:=UOWHF_Result[8] + 667400021+UOWHF_Add_c;
   		UOWHF_Add_c.8:=UOWHF_Result[8].31;
   		UOWHF_Result[8].31:=0;
   	End_If;
   	If UOWHF_Msg[3].[7] Then
   		UOWHF_Result[0]:=UOWHF_Result[0] + 615022266+UOWHF_Add_c;
   		UOWHF_Add_c.0:=UOWHF_Result[0].31;
   		UOWHF_Result[0].31:=0;
   		UOWHF_Result[1]:=UOWHF_Result[1] + 417783914+UOWHF_Add_c;
   		UOWHF_Add_c.1:=UOWHF_Result[1].31;
   		UOWHF_Result[1].31:=0;
   		UOWHF_Result[2]:=UOWHF_Result[2] + 359855697+UOWHF_Add_c;
   		UOWHF_Add_c.2:=UOWHF_Result[2].31;
   		UOWHF_Result[2].31:=0;
   		UOWHF_Result[3]:=UOWHF_Result[3] + 1256226964+UOWHF_Add_c;
   		UOWHF_Add_c.3:=UOWHF_Result[3].31;
   		UOWHF_Result[3].31:=0;
   		UOWHF_Result[4]:=UOWHF_Result[4] + 1440140153+UOWHF_Add_c;
   		UOWHF_Add_c.4:=UOWHF_Result[4].31;
   		UOWHF_Result[4].31:=0;
   		UOWHF_Result[5]:=UOWHF_Result[5] + 338797773+UOWHF_Add_c;
   		UOWHF_Add_c.5:=UOWHF_Result[5].31;
   		UOWHF_Result[5].31:=0;
   		UOWHF_Result[6]:=UOWHF_Result[6] + 1010450096+UOWHF_Add_c;
   		UOWHF_Add_c.6:=UOWHF_Result[6].31;
   		UOWHF_Result[6].31:=0;
   		UOWHF_Result[7]:=UOWHF_Result[7] + 194401209+UOWHF_Add_c;
   		UOWHF_Add_c.7:=UOWHF_Result[7].31;
   		UOWHF_Result[7].31:=0;
   		UOWHF_Result[8]:=UOWHF_Result[8] + 1421489120+UOWHF_Add_c;
   		UOWHF_Add_c.8:=UOWHF_Result[8].31;
   		UOWHF_Result[8].31:=0;
   	End_If;
   	If UOWHF_Msg[3].[8] Then
   		UOWHF_Result[0]:=UOWHF_Result[0] + 1456332546+UOWHF_Add_c;
   		UOWHF_Add_c.0:=UOWHF_Result[0].31;
   		UOWHF_Result[0].31:=0;
   		UOWHF_Result[1]:=UOWHF_Result[1] + 975978587+UOWHF_Add_c;
   		UOWHF_Add_c.1:=UOWHF_Result[1].31;
   		UOWHF_Result[1].31:=0;
   		UOWHF_Result[2]:=UOWHF_Result[2] + 297975624+UOWHF_Add_c;
   		UOWHF_Add_c.2:=UOWHF_Result[2].31;
   		UOWHF_Result[2].31:=0;
   		UOWHF_Result[3]:=UOWHF_Result[3] + 1138150841+UOWHF_Add_c;
   		UOWHF_Add_c.3:=UOWHF_Result[3].31;
   		UOWHF_Result[3].31:=0;
   		UOWHF_Result[4]:=UOWHF_Result[4] + 716758753+UOWHF_Add_c;
   		UOWHF_Add_c.4:=UOWHF_Result[4].31;
   		UOWHF_Result[4].31:=0;
   		UOWHF_Result[5]:=UOWHF_Result[5] + 1031342749+UOWHF_Add_c;
   		UOWHF_Add_c.5:=UOWHF_Result[5].31;
   		UOWHF_Result[5].31:=0;
   		UOWHF_Result[6]:=UOWHF_Result[6] + 1839835963+UOWHF_Add_c;
   		UOWHF_Add_c.6:=UOWHF_Result[6].31;
   		UOWHF_Result[6].31:=0;
   		UOWHF_Result[7]:=UOWHF_Result[7] + 2121125821+UOWHF_Add_c;
   		UOWHF_Add_c.7:=UOWHF_Result[7].31;
   		UOWHF_Result[7].31:=0;
   		UOWHF_Result[8]:=UOWHF_Result[8] + 59249464+UOWHF_Add_c;
   		UOWHF_Add_c.8:=UOWHF_Result[8].31;
   		UOWHF_Result[8].31:=0;
   	End_If;
   	If UOWHF_Msg[3].[9] Then
   		UOWHF_Result[0]:=UOWHF_Result[0] + 608589310+UOWHF_Add_c;
   		UOWHF_Add_c.0:=UOWHF_Result[0].31;
   		UOWHF_Result[0].31:=0;
   		UOWHF_Result[1]:=UOWHF_Result[1] + 222747636+UOWHF_Add_c;
   		UOWHF_Add_c.1:=UOWHF_Result[1].31;
   		UOWHF_Result[1].31:=0;
   		UOWHF_Result[2]:=UOWHF_Result[2] + 1937217872+UOWHF_Add_c;
   		UOWHF_Add_c.2:=UOWHF_Result[2].31;
   		UOWHF_Result[2].31:=0;
   		UOWHF_Result[3]:=UOWHF_Result[3] + 891453261+UOWHF_Add_c;
   		UOWHF_Add_c.3:=UOWHF_Result[3].31;
   		UOWHF_Result[3].31:=0;
   		UOWHF_Result[4]:=UOWHF_Result[4] + 13238587+UOWHF_Add_c;
   		UOWHF_Add_c.4:=UOWHF_Result[4].31;
   		UOWHF_Result[4].31:=0;
   		UOWHF_Result[5]:=UOWHF_Result[5] + 1969454841+UOWHF_Add_c;
   		UOWHF_Add_c.5:=UOWHF_Result[5].31;
   		UOWHF_Result[5].31:=0;
   		UOWHF_Result[6]:=UOWHF_Result[6] + 1376237148+UOWHF_Add_c;
   		UOWHF_Add_c.6:=UOWHF_Result[6].31;
   		UOWHF_Result[6].31:=0;
   		UOWHF_Result[7]:=UOWHF_Result[7] + 141767791+UOWHF_Add_c;
   		UOWHF_Add_c.7:=UOWHF_Result[7].31;
   		UOWHF_Result[7].31:=0;
   		UOWHF_Result[8]:=UOWHF_Result[8] + 507536491+UOWHF_Add_c;
   		UOWHF_Add_c.8:=UOWHF_Result[8].31;
   		UOWHF_Result[8].31:=0;
   	End_If;
   	If UOWHF_Msg[3].[10] Then
   		UOWHF_Result[0]:=UOWHF_Result[0] + 974915433+UOWHF_Add_c;
   		UOWHF_Add_c.0:=UOWHF_Result[0].31;
   		UOWHF_Result[0].31:=0;
   		UOWHF_Result[1]:=UOWHF_Result[1] + 1261907612+UOWHF_Add_c;
   		UOWHF_Add_c.1:=UOWHF_Result[1].31;
   		UOWHF_Result[1].31:=0;
   		UOWHF_Result[2]:=UOWHF_Result[2] + 1396568318+UOWHF_Add_c;
   		UOWHF_Add_c.2:=UOWHF_Result[2].31;
   		UOWHF_Result[2].31:=0;
   		UOWHF_Result[3]:=UOWHF_Result[3] + 2130031785+UOWHF_Add_c;
   		UOWHF_Add_c.3:=UOWHF_Result[3].31;
   		UOWHF_Result[3].31:=0;
   		UOWHF_Result[4]:=UOWHF_Result[4] + 1095665589+UOWHF_Add_c;
   		UOWHF_Add_c.4:=UOWHF_Result[4].31;
   		UOWHF_Result[4].31:=0;
   		UOWHF_Result[5]:=UOWHF_Result[5] + 372618186+UOWHF_Add_c;
   		UOWHF_Add_c.5:=UOWHF_Result[5].31;
   		UOWHF_Result[5].31:=0;
   		UOWHF_Result[6]:=UOWHF_Result[6] + 1004542979+UOWHF_Add_c;
   		UOWHF_Add_c.6:=UOWHF_Result[6].31;
   		UOWHF_Result[6].31:=0;
   		UOWHF_Result[7]:=UOWHF_Result[7] + 575139494+UOWHF_Add_c;
   		UOWHF_Add_c.7:=UOWHF_Result[7].31;
   		UOWHF_Result[7].31:=0;
   		UOWHF_Result[8]:=UOWHF_Result[8] + 1593362771+UOWHF_Add_c;
   		UOWHF_Add_c.8:=UOWHF_Result[8].31;
   		UOWHF_Result[8].31:=0;
   	End_If;
   	If UOWHF_Msg[3].[11] Then
   		UOWHF_Result[0]:=UOWHF_Result[0] + 1389992651+UOWHF_Add_c;
   		UOWHF_Add_c.0:=UOWHF_Result[0].31;
   		UOWHF_Result[0].31:=0;
   		UOWHF_Result[1]:=UOWHF_Result[1] + 474352379+UOWHF_Add_c;
   		UOWHF_Add_c.1:=UOWHF_Result[1].31;
   		UOWHF_Result[1].31:=0;
   		UOWHF_Result[2]:=UOWHF_Result[2] + 1567468459+UOWHF_Add_c;
   		UOWHF_Add_c.2:=UOWHF_Result[2].31;
   		UOWHF_Result[2].31:=0;
   		UOWHF_Result[3]:=UOWHF_Result[3] + 964686829+UOWHF_Add_c;
   		UOWHF_Add_c.3:=UOWHF_Result[3].31;
   		UOWHF_Result[3].31:=0;
   		UOWHF_Result[4]:=UOWHF_Result[4] + 1448886845+UOWHF_Add_c;
   		UOWHF_Add_c.4:=UOWHF_Result[4].31;
   		UOWHF_Result[4].31:=0;
   		UOWHF_Result[5]:=UOWHF_Result[5] + 1758603101+UOWHF_Add_c;